   t[5058] := 0;
   t[5059] := 0;
   t[5060] := 0;
   t[5061] := 0;
   t[5062] := 0;
   t[5063] := 0;
   t[5064] := 0;
   t[5065] := 0;
   t[5066] := 0;
   t[5067] := 0;
   t[5068] := 0;
   t[5069] := 0;
   t[5070] := 0;
   t[5071] := 0;
   t[5072] := 0;
   t[5073] := 0;
   t[5074] := 0;
   t[5075] := 0;
   t[5076] := 0;
   t[5077] := 0;
   t[5078] := 0;
   t[5079] := 0;
   t[5080] := 0;
   t[5081] := 0;
   t[5082] := 0;
   t[5083] := 0;
   t[5084] := 0;
   t[5085] := 0;
   t[5086] := 0;
   t[5087] := 0;
   t[5088] := 0;
   t[5089] := 0;
   t[5090] := 0;
   t[5091] := 0;
   t[5092] := 0;
   t[5093] := 0;
   t[5094] := 0;
   t[5095] := 0;
   t[5096] := 0;
   t[5097] := 0;
   t[5098] := 0;
   t[5099] := 0;
   t[5100] := 0;
   t[5101] := 0;
   t[5102] := 0;
   t[5103] := 0;
   t[5104] := 0;
   t[5105] := 0;
   t[5106] := 0;
   t[5107] := 0;
   t[5108] := 0;
   t[5109] := 0;
   t[5110] := 0;
   t[5111] := 0;
   t[5112] := 0;
   t[5113] := 0;
   t[5114] := 0;
   t[5115] := 0;
   t[5116] := 0;
   t[5117] := 0;
   t[5118] := 0;
   t[5119] := 0;
   t[5120] := 0;
   t[5121] := 0;
   t[5122] := 0;
   t[5123] := 0;
   t[5124] := 0;
   t[5125] := 0;
   t[5126] := 0;
   t[5127] := 0;
   t[5128] := 0;
   t[5129] := 0;
   t[5130] := 0;
   t[5131] := 0;
   t[5132] := 0;
   t[5133] := 0;
   t[5134] := 0;
   t[5135] := 0;
   t[5136] := 0;
   t[5137] := 0;
   t[5138] := 0;
   t[5139] := 0;
   t[5140] := 0;
   t[5141] := 0;
   t[5142] := 0;
   t[5143] := 0;
   t[5144] := 0;
   t[5145] := 0;
   t[5146] := 0;
   t[5147] := 0;
   t[5148] := 0;
   t[5149] := 0;
   t[5150] := 0;
   t[5151] := 0;
   t[5152] := 0;
   t[5153] := 0;
   t[5154] := 0;
   t[5155] := 0;
   t[5156] := 0;
   t[5157] := 0;
   t[5158] := 0;
   t[5159] := 0;
   t[5160] := 0;
   t[5161] := 0;
   t[5162] := 0;
   t[5163] := 0;
   t[5164] := 0;
   t[5165] := 0;
   t[5166] := 0;
   t[5167] := 0;
   t[5168] := 0;
   t[5169] := 0;
   t[5170] := 0;
   t[5171] := 0;
   t[5172] := 0;
   t[5173] := 0;
   t[5174] := 0;
   t[5175] := 0;
   t[5176] := 0;
   t[5177] := 0;
   t[5178] := 0;
   t[5179] := 0;
   t[5180] := 0;
   t[5181] := 0;
   t[5182] := 0;
   t[5183] := 0;
   t[5184] := 0;
   t[5185] := 0;
   t[5186] := 0;
   t[5187] := 0;
   t[5188] := 0;
   t[5189] := 0;
   t[5190] := 0;
   t[5191] := 0;
   t[5192] := 0;
   t[5193] := 0;
   t[5194] := 0;
   t[5195] := 0;
   t[5196] := 0;
   t[5197] := 0;
   t[5198] := 0;
   t[5199] := 0;
   t[5200] := 0;
   t[5201] := 0;
   t[5202] := 0;
   t[5203] := 0;
   t[5204] := 0;
   t[5205] := 0;
   t[5206] := 0;
   t[5207] := 0;
   t[5208] := 0;
   t[5209] := 0;
   t[5210] := 0;
   t[5211] := 0;
   t[5212] := 0;
   t[5213] := 0;
   t[5214] := 0;
   t[5215] := 0;
   t[5216] := 0;
   t[5217] := 0;
   t[5218] := 0;
   t[5219] := 0;
   t[5220] := 0;
   t[5221] := 0;
   t[5222] := 0;
   t[5223] := 0;
   t[5224] := 0;
   t[5225] := 0;
   t[5226] := 0;
   t[5227] := 0;
   t[5228] := 0;
   t[5229] := 0;
   t[5230] := 0;
   t[5231] := 0;
   t[5232] := 0;
   t[5233] := 0;
   t[5234] := 0;
   t[5235] := 0;
   t[5236] := 0;
   t[5237] := 0;
   t[5238] := 0;
   t[5239] := 0;
   t[5240] := 0;
   t[5241] := 0;
   t[5242] := 0;
   t[5243] := 0;
   t[5244] := 0;
   t[5245] := 0;
   t[5246] := 0;
   t[5247] := 0;
   t[5248] := 0;
   t[5249] := 0;
   t[5250] := 0;
   t[5251] := 0;
   t[5252] := 0;
   t[5253] := 0;
   t[5254] := 0;
   t[5255] := 0;
   t[5256] := 0;
   t[5257] := 0;
   t[5258] := 0;
   t[5259] := 0;
   t[5260] := 0;
   t[5261] := 0;
   t[5262] := 0;
   t[5263] := 0;
   t[5264] := 0;
   t[5265] := 0;
   t[5266] := 0;
   t[5267] := 0;
   t[5268] := 0;
   t[5269] := 0;
   t[5270] := 0;
   t[5271] := 0;
   t[5272] := 0;
   t[5273] := 0;
   t[5274] := 0;
   t[5275] := 0;
   t[5276] := 0;
   t[5277] := 0;
   t[5278] := 0;
   t[5279] := 0;
   t[5280] := 0;
   t[5281] := 0;
   t[5282] := 0;
   t[5283] := 0;
   t[5284] := 0;
   t[5285] := 0;
   t[5286] := 0;
   t[5287] := 0;
   t[5288] := 0;
   t[5289] := 0;
   t[5290] := 0;
   t[5291] := 0;
   t[5292] := 0;
   t[5293] := 0;
   t[5294] := 0;
   t[5295] := 0;
   t[5296] := 0;
   t[5297] := 0;
   t[5298] := 0;
   t[5299] := 0;
   t[5300] := 0;
   t[5301] := 0;
   t[5302] := 0;
   t[5303] := 0;
   t[5304] := 0;
   t[5305] := 0;
   t[5306] := 0;
   t[5307] := 0;
   t[5308] := 0;
   t[5309] := 0;
   t[5310] := 0;
   t[5311] := 0;
   t[5312] := 0;
   t[5313] := 0;
   t[5314] := 0;
   t[5315] := 0;
   t[5316] := 0;
   t[5317] := 0;
   t[5318] := 0;
   t[5319] := 0;
   t[5320] := 0;
   t[5321] := 0;
   t[5322] := 0;
   t[5323] := 0;
   t[5324] := 0;
   t[5325] := 0;
   t[5326] := 0;
   t[5327] := 0;
   t[5328] := 0;
   t[5329] := 0;
   t[5330] := 0;
   t[5331] := 0;
   t[5332] := 0;
   t[5333] := 0;
   t[5334] := 0;
   t[5335] := 0;
   t[5336] := 0;
   t[5337] := 0;
   t[5338] := 0;
   t[5339] := 0;
   t[5340] := 0;
   t[5341] := 0;
   t[5342] := 0;
   t[5343] := 0;
   t[5344] := 0;
   t[5345] := 0;
   t[5346] := 0;
   t[5347] := 0;
   t[5348] := 0;
   t[5349] := 0;
   t[5350] := 0;
   t[5351] := 0;
   t[5352] := 0;
   t[5353] := 0;
   t[5354] := 0;
   t[5355] := 0;
   t[5356] := 0;
   t[5357] := 0;
   t[5358] := 0;
   t[5359] := 0;
   t[5360] := 0;
   t[5361] := 0;
   t[5362] := 0;
   t[5363] := 0;
   t[5364] := 0;
   t[5365] := 0;
   t[5366] := 0;
   t[5367] := 0;
   t[5368] := 0;
   t[5369] := 0;
   t[5370] := 0;
   t[5371] := 0;
   t[5372] := 0;
   t[5373] := 0;
   t[5374] := 0;
   t[5375] := 0;
   t[5376] := 0;
   t[5377] := 0;
   t[5378] := 0;
   t[5379] := 0;
   t[5380] := 0;
   t[5381] := 0;
   t[5382] := 0;
   t[5383] := 0;
   t[5384] := 0;
   t[5385] := 0;
   t[5386] := 0;
   t[5387] := 0;
   t[5388] := 0;
   t[5389] := 0;
   t[5390] := 0;
   t[5391] := 0;
   t[5392] := 0;
   t[5393] := 0;
   t[5394] := 0;
   t[5395] := 0;
   t[5396] := 0;
   t[5397] := 0;
   t[5398] := 0;
   t[5399] := 0;
   t[5400] := 0;
   t[5401] := 0;
   t[5402] := 0;
   t[5403] := 0;
   t[5404] := 0;
   t[5405] := 0;
   t[5406] := 0;
   t[5407] := 0;
   t[5408] := 0;
   t[5409] := 0;
   t[5410] := 0;
   t[5411] := 0;
   t[5412] := 0;
   t[5413] := 0;
   t[5414] := 0;
   t[5415] := 0;
   t[5416] := 0;
   t[5417] := 0;
   t[5418] := 0;
   t[5419] := 0;
   t[5420] := 0;
   t[5421] := 0;
   t[5422] := 0;
   t[5423] := 0;
   t[5424] := 0;
   t[5425] := 0;
   t[5426] := 0;
   t[5427] := 0;
   t[5428] := 0;
   t[5429] := 0;
   t[5430] := 0;
   t[5431] := 0;
   t[5432] := 0;
   t[5433] := 0;
   t[5434] := 0;
   t[5435] := 0;
   t[5436] := 0;
   t[5437] := 0;
   t[5438] := 0;
   t[5439] := 0;
   t[5440] := 0;
   t[5441] := 0;
   t[5442] := 0;
   t[5443] := 0;
   t[5444] := 0;
   t[5445] := 0;
   t[5446] := 0;
   t[5447] := 0;
   t[5448] := 0;
   t[5449] := 0;
   t[5450] := 0;
   t[5451] := 0;
   t[5452] := 0;
   t[5453] := 0;
   t[5454] := 0;
   t[5455] := 0;
   t[5456] := 0;
   t[5457] := 0;
   t[5458] := 0;
   t[5459] := 0;
   t[5460] := 0;
   t[5461] := 0;
   t[5462] := 0;
   t[5463] := 0;
   t[5464] := 0;
   t[5465] := 0;
   t[5466] := 0;
   t[5467] := 0;
   t[5468] := 0;
   t[5469] := 0;
   t[5470] := 0;
   t[5471] := 0;
   t[5472] := 0;
   t[5473] := 0;
   t[5474] := 0;
   t[5475] := 0;
   t[5476] := 0;
   t[5477] := 0;
   t[5478] := 0;
   t[5479] := 0;
   t[5480] := 0;
   t[5481] := 0;
   t[5482] := 0;
   t[5483] := 0;
   t[5484] := 0;
   t[5485] := 0;
   t[5486] := 0;
   t[5487] := 0;
   t[5488] := 0;
   t[5489] := 0;
   t[5490] := 0;
   t[5491] := 0;
   t[5492] := 0;
   t[5493] := 0;
   t[5494] := 0;
   t[5495] := 0;
   t[5496] := 0;
   t[5497] := 0;
   t[5498] := 0;
   t[5499] := 0;
   t[5500] := 0;
   t[5501] := 0;
   t[5502] := 0;
   t[5503] := 0;
   t[5504] := 0;
   t[5505] := 0;
   t[5506] := 0;
   t[5507] := 0;
   t[5508] := 0;
   t[5509] := 0;
   t[5510] := 0;
   t[5511] := 0;
   t[5512] := 0;
   t[5513] := 0;
   t[5514] := 0;
   t[5515] := 0;
   t[5516] := 0;
   t[5517] := 0;
   t[5518] := 0;
   t[5519] := 0;
   t[5520] := 0;
   t[5521] := 0;
   t[5522] := 0;
   t[5523] := 0;
   t[5524] := 0;
   t[5525] := 0;
   t[5526] := 0;
   t[5527] := 0;
   t[5528] := 0;
   t[5529] := 0;
   t[5530] := 0;
   t[5531] := 0;
   t[5532] := 0;
   t[5533] := 0;
   t[5534] := 0;
   t[5535] := 0;
   t[5536] := 0;
   t[5537] := 0;
   t[5538] := 0;
   t[5539] := 0;
   t[5540] := 0;
   t[5541] := 0;
   t[5542] := 0;
   t[5543] := 0;
   t[5544] := 0;
   t[5545] := 0;
   t[5546] := 0;
   t[5547] := 0;
   t[5548] := 0;
   t[5549] := 0;
   t[5550] := 0;
   t[5551] := 0;
   t[5552] := 0;
   t[5553] := 0;
   t[5554] := 0;
   t[5555] := 0;
   t[5556] := 0;
   t[5557] := 0;
   t[5558] := 0;
   t[5559] := 0;
   t[5560] := 0;
   t[5561] := 0;
   t[5562] := 0;
   t[5563] := 0;
   t[5564] := 0;
   t[5565] := 0;
   t[5566] := 0;
   t[5567] := 0;
   t[5568] := 0;
   t[5569] := 0;
   t[5570] := 0;
   t[5571] := 0;
   t[5572] := 0;
   t[5573] := 0;
   t[5574] := 0;
   t[5575] := 0;
   t[5576] := 0;
   t[5577] := 0;
   t[5578] := 0;
   t[5579] := 0;
   t[5580] := 0;
   t[5581] := 0;
   t[5582] := 0;
   t[5583] := 0;
   t[5584] := 0;
   t[5585] := 0;
   t[5586] := 0;
   t[5587] := 0;
   t[5588] := 0;
   t[5589] := 0;
   t[5590] := 0;
   t[5591] := 0;
   t[5592] := 0;
   t[5593] := 0;
   t[5594] := 0;
   t[5595] := 0;
   t[5596] := 0;
   t[5597] := 0;
   t[5598] := 0;
   t[5599] := 0;
   t[5600] := 0;
   t[5601] := 0;
   t[5602] := 0;
   t[5603] := 0;
   t[5604] := 0;
   t[5605] := 0;
   t[5606] := 0;
   t[5607] := 0;
   t[5608] := 0;
   t[5609] := 0;
   t[5610] := 0;
   t[5611] := 0;
   t[5612] := 0;
   t[5613] := 0;
   t[5614] := 0;
   t[5615] := 0;
   t[5616] := 0;
   t[5617] := 0;
   t[5618] := 0;
   t[5619] := 0;
   t[5620] := 0;
   t[5621] := 0;
   t[5622] := 0;
   t[5623] := 0;
   t[5624] := 0;
   t[5625] := 0;
   t[5626] := 0;
   t[5627] := 0;
   t[5628] := 0;
   t[5629] := 0;
   t[5630] := 0;
   t[5631] := 0;
   t[5632] := 0;
   t[5633] := 0;
   t[5634] := 0;
   t[5635] := 0;
   t[5636] := 0;
   t[5637] := 0;
   t[5638] := 0;
   t[5639] := 0;
   t[5640] := 0;
   t[5641] := 0;
   t[5642] := 0;
   t[5643] := 0;
   t[5644] := 0;
   t[5645] := 0;
   t[5646] := 0;
   t[5647] := 0;
   t[5648] := 0;
   t[5649] := 0;
   t[5650] := 0;
   t[5651] := 0;
   t[5652] := 0;
   t[5653] := 0;
   t[5654] := 0;
   t[5655] := 0;
   t[5656] := 0;
   t[5657] := 0;
   t[5658] := 0;
   t[5659] := 0;
   t[5660] := 0;
   t[5661] := 0;
   t[5662] := 0;
   t[5663] := 0;
   t[5664] := 0;
   t[5665] := 0;
   t[5666] := 0;
   t[5667] := 0;
   t[5668] := 0;
   t[5669] := 0;
   t[5670] := 0;
   t[5671] := 0;
   t[5672] := 0;
   t[5673] := 0;
   t[5674] := 0;
   t[5675] := 0;
   t[5676] := 0;
   t[5677] := 0;
   t[5678] := 0;
   t[5679] := 0;
   t[5680] := 0;
   t[5681] := 0;
   t[5682] := 0;
   t[5683] := 0;
   t[5684] := 0;
   t[5685] := 0;
   t[5686] := 0;
   t[5687] := 0;
   t[5688] := 0;
   t[5689] := 0;
   t[5690] := 0;
   t[5691] := 0;
   t[5692] := 0;
   t[5693] := 0;
   t[5694] := 0;
   t[5695] := 0;
   t[5696] := 0;
   t[5697] := 0;
   t[5698] := 0;
   t[5699] := 0;
   t[5700] := 0;
   t[5701] := 0;
   t[5702] := 0;
   t[5703] := 0;
   t[5704] := 0;
   t[5705] := 0;
   t[5706] := 0;
   t[5707] := 0;
   t[5708] := 0;
   t[5709] := 0;
   t[5710] := 0;
   t[5711] := 0;
   t[5712] := 0;
   t[5713] := 0;
   t[5714] := 0;
   t[5715] := 0;
   t[5716] := 0;
   t[5717] := 0;
   t[5718] := 0;
   t[5719] := 0;
   t[5720] := 0;
   t[5721] := 0;
   t[5722] := 0;
   t[5723] := 0;
   t[5724] := 0;
   t[5725] := 0;
   t[5726] := 0;
   t[5727] := 0;
   t[5728] := 0;
   t[5729] := 0;
   t[5730] := 0;
   t[5731] := 0;
   t[5732] := 0;
   t[5733] := 0;
   t[5734] := 0;
   t[5735] := 0;
   t[5736] := 0;
   t[5737] := 0;
   t[5738] := 0;
   t[5739] := 0;
   t[5740] := 0;
   t[5741] := 0;
   t[5742] := 0;
   t[5743] := 0;
   t[5744] := 0;
   t[5745] := 0;
   t[5746] := 0;
   t[5747] := 0;
   t[5748] := 0;
   t[5749] := 0;
   t[5750] := 0;
   t[5751] := 0;
   t[5752] := 0;
   t[5753] := 0;
   t[5754] := 0;
   t[5755] := 0;
   t[5756] := 0;
   t[5757] := 0;
   t[5758] := 0;
   t[5759] := 0;
   t[5760] := 0;
   t[5761] := 0;
   t[5762] := 0;
   t[5763] := 0;
   t[5764] := 0;
   t[5765] := 0;
   t[5766] := 0;
   t[5767] := 0;
   t[5768] := 0;
   t[5769] := 0;
   t[5770] := 0;
   t[5771] := 0;
   t[5772] := 0;
   t[5773] := 0;
   t[5774] := 0;
   t[5775] := 0;
   t[5776] := 0;
   t[5777] := 0;
   t[5778] := 0;
   t[5779] := 0;
   t[5780] := 0;
   t[5781] := 0;
   t[5782] := 0;
   t[5783] := 0;
   t[5784] := 0;
   t[5785] := 0;
   t[5786] := 0;
   t[5787] := 0;
   t[5788] := 0;
   t[5789] := 0;
   t[5790] := 0;
   t[5791] := 0;
   t[5792] := 0;
   t[5793] := 0;
   t[5794] := 0;
   t[5795] := 0;
   t[5796] := 0;
   t[5797] := 0;
   t[5798] := 0;
   t[5799] := 0;
   t[5800] := 0;
   t[5801] := 0;
   t[5802] := 0;
   t[5803] := 0;
   t[5804] := 0;
   t[5805] := 0;
   t[5806] := 0;
   t[5807] := 0;
   t[5808] := 0;
   t[5809] := 0;
   t[5810] := 0;
   t[5811] := 0;
   t[5812] := 0;
   t[5813] := 0;
   t[5814] := 0;
   t[5815] := 0;
   t[5816] := 0;
   t[5817] := 0;
   t[5818] := 0;
   t[5819] := 0;
   t[5820] := 0;
   t[5821] := 0;
   t[5822] := 0;
   t[5823] := 0;
   t[5824] := 0;
   t[5825] := 0;
   t[5826] := 0;
   t[5827] := 0;
   t[5828] := 0;
   t[5829] := 0;
   t[5830] := 0;
   t[5831] := 0;
   t[5832] := 0;
   t[5833] := 0;
   t[5834] := 0;
   t[5835] := 0;
   t[5836] := 0;
   t[5837] := 0;
   t[5838] := 0;
   t[5839] := 0;
   t[5840] := 0;
   t[5841] := 0;
   t[5842] := 0;
   t[5843] := 0;
   t[5844] := 0;
   t[5845] := 0;
   t[5846] := 0;
   t[5847] := 0;
   t[5848] := 0;
   t[5849] := 0;
   t[5850] := 0;
   t[5851] := 0;
   t[5852] := 0;
   t[5853] := 0;
   t[5854] := 0;
   t[5855] := 0;
   t[5856] := 0;
   t[5857] := 0;
   t[5858] := 0;
   t[5859] := 0;
   t[5860] := 0;
   t[5861] := 0;
   t[5862] := 0;
   t[5863] := 0;
   t[5864] := 0;
   t[5865] := 0;
   t[5866] := 0;
   t[5867] := 0;
   t[5868] := 0;
   t[5869] := 0;
   t[5870] := 0;
   t[5871] := 0;
   t[5872] := 0;
   t[5873] := 0;
   t[5874] := 0;
   t[5875] := 0;
   t[5876] := 0;
   t[5877] := 0;
   t[5878] := 0;
   t[5879] := 0;
   t[5880] := 0;
   t[5881] := 0;
   t[5882] := 0;
   t[5883] := 0;
   t[5884] := 0;
   t[5885] := 0;
   t[5886] := 0;
   t[5887] := 0;
   t[5888] := 0;
   t[5889] := 0;
   t[5890] := 0;
   t[5891] := 0;
   t[5892] := 0;
   t[5893] := 0;
   t[5894] := 0;
   t[5895] := 0;
   t[5896] := 0;
   t[5897] := 0;
   t[5898] := 0;
   t[5899] := 0;
   t[5900] := 0;
   t[5901] := 0;
   t[5902] := 0;
   t[5903] := 0;
   t[5904] := 0;
   t[5905] := 0;
   t[5906] := 0;
   t[5907] := 0;
   t[5908] := 0;
   t[5909] := 0;
   t[5910] := 0;
   t[5911] := 0;
   t[5912] := 0;
   t[5913] := 0;
   t[5914] := 0;
   t[5915] := 0;
   t[5916] := 0;
   t[5917] := 0;
   t[5918] := 0;
   t[5919] := 0;
   t[5920] := 0;
   t[5921] := 0;
   t[5922] := 0;
   t[5923] := 0;
   t[5924] := 0;
   t[5925] := 0;
   t[5926] := 0;
   t[5927] := 0;
   t[5928] := 0;
   t[5929] := 0;
   t[5930] := 0;
   t[5931] := 0;
   t[5932] := 0;
   t[5933] := 0;
   t[5934] := 0;
   t[5935] := 0;
   t[5936] := 0;
   t[5937] := 0;
   t[5938] := 0;
   t[5939] := 0;
   t[5940] := 0;
   t[5941] := 0;
   t[5942] := 0;
   t[5943] := 0;
   t[5944] := 0;
   t[5945] := 0;
   t[5946] := 0;
   t[5947] := 0;
   t[5948] := 0;
   t[5949] := 0;
   t[5950] := 0;
   t[5951] := 0;
   t[5952] := 0;
   t[5953] := 0;
   t[5954] := 0;
   t[5955] := 0;
   t[5956] := 0;
   t[5957] := 0;
   t[5958] := 0;
   t[5959] := 0;
   t[5960] := 0;
   t[5961] := 0;
   t[5962] := 0;
   t[5963] := 0;
   t[5964] := 0;
   t[5965] := 0;
   t[5966] := 0;
   t[5967] := 0;
   t[5968] := 0;
   t[5969] := 0;
   t[5970] := 0;
   t[5971] := 0;
   t[5972] := 0;
   t[5973] := 0;
   t[5974] := 0;
   t[5975] := 0;
   t[5976] := 0;
   t[5977] := 0;
   t[5978] := 0;
   t[5979] := 0;
   t[5980] := 0;
   t[5981] := 0;
   t[5982] := 0;
   t[5983] := 0;
   t[5984] := 0;
   t[5985] := 0;
   t[5986] := 0;
   t[5987] := 0;
   t[5988] := 0;
   t[5989] := 0;
   t[5990] := 0;
   t[5991] := 0;
   t[5992] := 0;
   t[5993] := 0;
   t[5994] := 0;
   t[5995] := 0;
   t[5996] := 0;
   t[5997] := 0;
   t[5998] := 0;
   t[5999] := 0;
   t[6000] := 0;
   t[6001] := 0;
   t[6002] := 0;
   t[6003] := 0;
   t[6004] := 0;
   t[6005] := 0;
   t[6006] := 0;
   t[6007] := 0;
   t[6008] := 0;
   t[6009] := 0;
   t[6010] := 0;
   t[6011] := 0;
   t[6012] := 0;
   t[6013] := 0;
   t[6014] := 0;
   t[6015] := 0;
   t[6016] := 0;
   t[6017] := 0;
   t[6018] := 0;
   t[6019] := 0;
   t[6020] := 0;
   t[6021] := 0;
   t[6022] := 0;
   t[6023] := 0;
   t[6024] := 0;
   t[6025] := 0;
   t[6026] := 0;
   t[6027] := 0;
   t[6028] := 0;
   t[6029] := 0;
   t[6030] := 0;
   t[6031] := 0;
   t[6032] := 0;
   t[6033] := 0;
   t[6034] := 0;
   t[6035] := 0;
   t[6036] := 0;
   t[6037] := 0;
   t[6038] := 0;
   t[6039] := 0;
   t[6040] := 0;
   t[6041] := 0;
   t[6042] := 0;
   t[6043] := 0;
   t[6044] := 0;
   t[6045] := 0;
   t[6046] := 0;
   t[6047] := 0;
   t[6048] := 0;
   t[6049] := 0;
   t[6050] := 0;
   t[6051] := 0;
   t[6052] := 0;
   t[6053] := 0;
   t[6054] := 0;
   t[6055] := 0;
   t[6056] := 0;
   t[6057] := 0;
   t[6058] := 0;
   t[6059] := 0;
   t[6060] := 0;
   t[6061] := 0;
   t[6062] := 0;
   t[6063] := 0;
   t[6064] := 0;
   t[6065] := 0;
   t[6066] := 0;
   t[6067] := 0;
   t[6068] := 0;
   t[6069] := 0;
   t[6070] := 0;
   t[6071] := 0;
   t[6072] := 0;
   t[6073] := 0;
   t[6074] := 0;
   t[6075] := 0;
   t[6076] := 0;
   t[6077] := 0;
   t[6078] := 0;
   t[6079] := 0;
   t[6080] := 0;
   t[6081] := 0;
   t[6082] := 0;
   t[6083] := 0;
   t[6084] := 0;
   t[6085] := 0;
   t[6086] := 0;
   t[6087] := 0;
   t[6088] := 0;
   t[6089] := 0;
   t[6090] := 0;
   t[6091] := 0;
   t[6092] := 0;
   t[6093] := 0;
   t[6094] := 0;
   t[6095] := 0;
   t[6096] := 0;
   t[6097] := 0;
   t[6098] := 0;
   t[6099] := 0;
   t[6100] := 0;
   t[6101] := 0;
   t[6102] := 0;
   t[6103] := 0;
   t[6104] := 0;
   t[6105] := 0;
   t[6106] := 0;
   t[6107] := 0;
   t[6108] := 0;
   t[6109] := 0;
   t[6110] := 0;
   t[6111] := 0;
   t[6112] := 0;
   t[6113] := 0;
   t[6114] := 0;
   t[6115] := 0;
   t[6116] := 0;
   t[6117] := 0;
   t[6118] := 0;
   t[6119] := 0;
   t[6120] := 0;
   t[6121] := 0;
   t[6122] := 0;
   t[6123] := 0;
   t[6124] := 0;
   t[6125] := 0;
   t[6126] := 0;
   t[6127] := 0;
   t[6128] := 0;
   t[6129] := 0;
   t[6130] := 0;
   t[6131] := 0;
   t[6132] := 0;
   t[6133] := 0;
   t[6134] := 0;
   t[6135] := 0;
   t[6136] := 0;
   t[6137] := 0;
   t[6138] := 0;
   t[6139] := 0;
   t[6140] := 0;
   t[6141] := 0;
   t[6142] := 0;
   t[6143] := 0;
   t[6144] := 0;
   t[6145] := 0;
   t[6146] := 0;
   t[6147] := 0;
   t[6148] := 0;
   t[6149] := 0;
   t[6150] := 0;
   t[6151] := 0;
   t[6152] := 0;
   t[6153] := 0;
   t[6154] := 0;
   t[6155] := 0;
   t[6156] := 0;
   t[6157] := 0;
   t[6158] := 0;
   t[6159] := 0;
   t[6160] := 0;
   t[6161] := 0;
   t[6162] := 0;
   t[6163] := 0;
   t[6164] := 0;
   t[6165] := 0;
   t[6166] := 0;
   t[6167] := 0;
   t[6168] := 0;
   t[6169] := 0;
   t[6170] := 0;
   t[6171] := 0;
   t[6172] := 0;
   t[6173] := 0;
   t[6174] := 0;
   t[6175] := 0;
   t[6176] := 0;
   t[6177] := 0;
   t[6178] := 0;
   t[6179] := 0;
   t[6180] := 0;
   t[6181] := 0;
   t[6182] := 0;
   t[6183] := 0;
   t[6184] := 0;
   t[6185] := 0;
   t[6186] := 0;
   t[6187] := 0;
   t[6188] := 0;
   t[6189] := 0;
   t[6190] := 0;
   t[6191] := 0;
   t[6192] := 0;
   t[6193] := 0;
   t[6194] := 0;
   t[6195] := 0;
   t[6196] := 0;
   t[6197] := 0;
   t[6198] := 0;
   t[6199] := 0;
   t[6200] := 0;
   t[6201] := 0;
   t[6202] := 0;
   t[6203] := 0;
   t[6204] := 0;
   t[6205] := 0;
   t[6206] := 0;
   t[6207] := 0;
   t[6208] := 0;
   t[6209] := 0;
   t[6210] := 0;
   t[6211] := 0;
   t[6212] := 0;
   t[6213] := 0;
   t[6214] := 0;
   t[6215] := 0;
   t[6216] := 0;
   t[6217] := 0;
   t[6218] := 0;
   t[6219] := 0;
   t[6220] := 0;
   t[6221] := 0;
   t[6222] := 0;
   t[6223] := 0;
   t[6224] := 0;
   t[6225] := 0;
   t[6226] := 0;
   t[6227] := 0;
   t[6228] := 0;
   t[6229] := 0;
   t[6230] := 0;
   t[6231] := 0;
   t[6232] := 0;
   t[6233] := 0;
   t[6234] := 0;
   t[6235] := 0;
   t[6236] := 0;
   t[6237] := 0;
   t[6238] := 0;
   t[6239] := 0;
   t[6240] := 0;
   t[6241] := 0;
   t[6242] := 0;
   t[6243] := 0;
   t[6244] := 0;
   t[6245] := 0;
   t[6246] := 0;
   t[6247] := 0;
   t[6248] := 0;
   t[6249] := 0;
   t[6250] := 0;
   t[6251] := 0;
   t[6252] := 0;
   t[6253] := 0;
   t[6254] := 0;
   t[6255] := 0;
   t[6256] := 0;
   t[6257] := 0;
   t[6258] := 0;
   t[6259] := 0;
   t[6260] := 0;
   t[6261] := 0;
   t[6262] := 0;
   t[6263] := 0;
   t[6264] := 0;
   t[6265] := 0;
   t[6266] := 0;
   t[6267] := 0;
   t[6268] := 0;
   t[6269] := 0;
   t[6270] := 0;
   t[6271] := 0;
   t[6272] := 0;
   t[6273] := 0;
   t[6274] := 0;
   t[6275] := 0;
   t[6276] := 0;
   t[6277] := 0;
   t[6278] := 0;
   t[6279] := 0;
   t[6280] := 0;
   t[6281] := 0;
   t[6282] := 0;
   t[6283] := 0;
   t[6284] := 0;
   t[6285] := 0;
   t[6286] := 0;
   t[6287] := 0;
   t[6288] := 0;
   t[6289] := 0;
   t[6290] := 0;
   t[6291] := 0;
   t[6292] := 0;
   t[6293] := 0;
   t[6294] := 0;
   t[6295] := 0;
   t[6296] := 0;
   t[6297] := 0;
   t[6298] := 0;
   t[6299] := 0;
   t[6300] := 0;
   t[6301] := 0;
   t[6302] := 0;
   t[6303] := 0;
   t[6304] := 0;
   t[6305] := 0;
   t[6306] := 0;
   t[6307] := 0;
   t[6308] := 0;
   t[6309] := 0;
   t[6310] := 0;
   t[6311] := 0;
   t[6312] := 0;
   t[6313] := 0;
   t[6314] := 0;
   t[6315] := 0;
   t[6316] := 0;
   t[6317] := 0;
   t[6318] := 0;
   t[6319] := 0;
   t[6320] := 0;
   t[6321] := 0;
   t[6322] := 0;
   t[6323] := 0;
   t[6324] := 0;
   t[6325] := 0;
   t[6326] := 0;
   t[6327] := 0;
   t[6328] := 0;
   t[6329] := 0;
   t[6330] := 0;
   t[6331] := 0;
   t[6332] := 0;
   t[6333] := 0;
   t[6334] := 0;
   t[6335] := 0;
   t[6336] := 0;
   t[6337] := 0;
   t[6338] := 0;
   t[6339] := 0;
   t[6340] := 0;
   t[6341] := 0;
   t[6342] := 0;
   t[6343] := 0;
   t[6344] := 0;
   t[6345] := 0;
   t[6346] := 0;
   t[6347] := 0;
   t[6348] := 0;
   t[6349] := 0;
   t[6350] := 0;
   t[6351] := 0;
   t[6352] := 0;
   t[6353] := 0;
   t[6354] := 0;
   t[6355] := 0;
   t[6356] := 0;
   t[6357] := 0;
   t[6358] := 0;
   t[6359] := 0;
   t[6360] := 0;
   t[6361] := 0;
   t[6362] := 0;
   t[6363] := 0;
   t[6364] := 0;
   t[6365] := 0;
   t[6366] := 0;
   t[6367] := 0;
   t[6368] := 0;
   t[6369] := 0;
   t[6370] := 0;
   t[6371] := 0;
   t[6372] := 0;
   t[6373] := 0;
   t[6374] := 0;
   t[6375] := 0;
   t[6376] := 0;
   t[6377] := 0;
   t[6378] := 0;
   t[6379] := 0;
   t[6380] := 0;
   t[6381] := 0;
   t[6382] := 0;
   t[6383] := 0;
   t[6384] := 0;
   t[6385] := 0;
   t[6386] := 0;
   t[6387] := 0;
   t[6388] := 0;
   t[6389] := 0;
   t[6390] := 0;
   t[6391] := 0;
   t[6392] := 0;
   t[6393] := 0;
   t[6394] := 0;
   t[6395] := 0;
   t[6396] := 0;
   t[6397] := 0;
   t[6398] := 0;
   t[6399] := 0;
   t[6400] := 0;
   t[6401] := 0;
   t[6402] := 0;
   t[6403] := 0;
   t[6404] := 0;
   t[6405] := 0;
   t[6406] := 0;
   t[6407] := 0;
   t[6408] := 0;
   t[6409] := 0;
   t[6410] := 0;
   t[6411] := 0;
   t[6412] := 0;
   t[6413] := 0;
   t[6414] := 0;
   t[6415] := 0;
   t[6416] := 0;
   t[6417] := 0;
   t[6418] := 0;
   t[6419] := 0;
   t[6420] := 0;
   t[6421] := 0;
   t[6422] := 0;
   t[6423] := 0;
   t[6424] := 0;
   t[6425] := 0;
   t[6426] := 0;
   t[6427] := 0;
   t[6428] := 0;
   t[6429] := 0;
   t[6430] := 0;
   t[6431] := 0;
   t[6432] := 0;
   t[6433] := 0;
   t[6434] := 0;
   t[6435] := 0;
   t[6436] := 0;
   t[6437] := 0;
   t[6438] := 0;
   t[6439] := 0;
   t[6440] := 0;
   t[6441] := 0;
   t[6442] := 0;
   t[6443] := 0;
   t[6444] := 0;
   t[6445] := 0;
   t[6446] := 0;
   t[6447] := 0;
   t[6448] := 0;
   t[6449] := 0;
   t[6450] := 0;
   t[6451] := 0;
   t[6452] := 0;
   t[6453] := 0;
   t[6454] := 0;
   t[6455] := 0;
   t[6456] := 0;
   t[6457] := 0;
   t[6458] := 0;
   t[6459] := 0;
   t[6460] := 0;
   t[6461] := 0;
   t[6462] := 0;
   t[6463] := 0;
   t[6464] := 0;
   t[6465] := 0;
   t[6466] := 0;
   t[6467] := 0;
   t[6468] := 0;
   t[6469] := 0;
   t[6470] := 0;
   t[6471] := 0;
   t[6472] := 0;
   t[6473] := 0;
   t[6474] := 0;
   t[6475] := 0;
   t[6476] := 0;
   t[6477] := 0;
   t[6478] := 0;
   t[6479] := 0;
   t[6480] := 0;
   t[6481] := 0;
   t[6482] := 0;
   t[6483] := 0;
   t[6484] := 0;
   t[6485] := 0;
   t[6486] := 0;
   t[6487] := 0;
   t[6488] := 0;
   t[6489] := 0;
   t[6490] := 0;
   t[6491] := 0;
   t[6492] := 0;
   t[6493] := 0;
   t[6494] := 0;
   t[6495] := 0;
   t[6496] := 0;
   t[6497] := 0;
   t[6498] := 0;
   t[6499] := 0;
   t[6500] := 0;
   t[6501] := 0;
   t[6502] := 0;
   t[6503] := 0;
   t[6504] := 0;
   t[6505] := 0;
   t[6506] := 0;
   t[6507] := 0;
   t[6508] := 0;
   t[6509] := 0;
   t[6510] := 0;
   t[6511] := 0;
   t[6512] := 0;
   t[6513] := 0;
   t[6514] := 0;
   t[6515] := 0;
   t[6516] := 0;
   t[6517] := 0;
   t[6518] := 0;
   t[6519] := 0;
   t[6520] := 0;
   t[6521] := 0;
   t[6522] := 0;
   t[6523] := 0;
   t[6524] := 0;
   t[6525] := 0;
   t[6526] := 0;
   t[6527] := 0;
   t[6528] := 0;
   t[6529] := 0;
   t[6530] := 0;
   t[6531] := 0;
   t[6532] := 0;
   t[6533] := 0;
   t[6534] := 0;
   t[6535] := 0;
   t[6536] := 0;
   t[6537] := 0;
   t[6538] := 0;
   t[6539] := 0;
   t[6540] := 0;
   t[6541] := 0;
   t[6542] := 0;
   t[6543] := 0;
   t[6544] := 0;
   t[6545] := 0;
   t[6546] := 0;
   t[6547] := 0;
   t[6548] := 0;
   t[6549] := 0;
   t[6550] := 0;
   t[6551] := 0;
   t[6552] := 0;
   t[6553] := 0;
   t[6554] := 0;
   t[6555] := 0;
   t[6556] := 0;
   t[6557] := 0;
   t[6558] := 0;
   t[6559] := 0;
   t[6560] := 0;
   t[6561] := 0;
   t[6562] := 0;
   t[6563] := 0;
   t[6564] := 0;
   t[6565] := 0;
   t[6566] := 0;
   t[6567] := 0;
   t[6568] := 0;
   t[6569] := 0;
   t[6570] := 0;
   t[6571] := 0;
   t[6572] := 0;
   t[6573] := 0;
   t[6574] := 0;
   t[6575] := 0;
   t[6576] := 0;
   t[6577] := 0;
   t[6578] := 0;
   t[6579] := 0;
   t[6580] := 0;
   t[6581] := 0;
   t[6582] := 0;
   t[6583] := 0;
   t[6584] := 0;
   t[6585] := 0;
   t[6586] := 0;
   t[6587] := 0;
   t[6588] := 0;
   t[6589] := 0;
   t[6590] := 0;
   t[6591] := 0;
   t[6592] := 0;
   t[6593] := 0;
   t[6594] := 0;
   t[6595] := 0;
   t[6596] := 0;
   t[6597] := 0;
   t[6598] := 0;
   t[6599] := 0;
   t[6600] := 0;
   t[6601] := 0;
   t[6602] := 0;
   t[6603] := 0;
   t[6604] := 0;
   t[6605] := 0;
   t[6606] := 0;
   t[6607] := 0;
   t[6608] := 0;
   t[6609] := 0;
   t[6610] := 0;
   t[6611] := 0;
   t[6612] := 0;
   t[6613] := 0;
   t[6614] := 0;
   t[6615] := 0;
   t[6616] := 0;
   t[6617] := 0;
   t[6618] := 0;
   t[6619] := 0;
   t[6620] := 0;
   t[6621] := 0;
   t[6622] := 0;
   t[6623] := 0;
   t[6624] := 0;
   t[6625] := 0;
   t[6626] := 0;
   t[6627] := 0;
   t[6628] := 0;
   t[6629] := 0;
   t[6630] := 0;
   t[6631] := 0;
   t[6632] := 0;
   t[6633] := 0;
   t[6634] := 0;
   t[6635] := 0;
   t[6636] := 0;
   t[6637] := 0;
   t[6638] := 0;
   t[6639] := 0;
   t[6640] := 0;
   t[6641] := 0;
   t[6642] := 0;
   t[6643] := 0;
   t[6644] := 0;
   t[6645] := 0;
   t[6646] := 0;
   t[6647] := 0;
   t[6648] := 0;
   t[6649] := 0;
   t[6650] := 0;
   t[6651] := 0;
   t[6652] := 0;
   t[6653] := 0;
   t[6654] := 0;
   t[6655] := 0;
   t[6656] := 0;
   t[6657] := 0;
   t[6658] := 0;
   t[6659] := 0;
   t[6660] := 0;
   t[6661] := 0;
   t[6662] := 0;
   t[6663] := 0;
   t[6664] := 0;
   t[6665] := 0;
   t[6666] := 0;
   t[6667] := 0;
   t[6668] := 0;
   t[6669] := 0;
   t[6670] := 0;
   t[6671] := 0;
   t[6672] := 0;
   t[6673] := 0;
   t[6674] := 0;
   t[6675] := 0;
   t[6676] := 0;
   t[6677] := 0;
   t[6678] := 0;
   t[6679] := 0;
   t[6680] := 0;
   t[6681] := 0;
   t[6682] := 0;
   t[6683] := 0;
   t[6684] := 0;
   t[6685] := 0;
   t[6686] := 0;
   t[6687] := 0;
   t[6688] := 0;
   t[6689] := 0;
   t[6690] := 0;
   t[6691] := 0;
   t[6692] := 0;
   t[6693] := 0;
   t[6694] := 0;
   t[6695] := 0;
   t[6696] := 0;
   t[6697] := 0;
   t[6698] := 0;
   t[6699] := 0;
   t[6700] := 0;
   t[6701] := 0;
   t[6702] := 0;
   t[6703] := 0;
   t[6704] := 0;
   t[6705] := 0;
   t[6706] := 0;
   t[6707] := 0;
   t[6708] := 0;
   t[6709] := 0;
   t[6710] := 0;
   t[6711] := 0;
   t[6712] := 0;
   t[6713] := 0;
   t[6714] := 0;
   t[6715] := 0;
   t[6716] := 0;
   t[6717] := 0;
   t[6718] := 0;
   t[6719] := 0;
   t[6720] := 0;
   t[6721] := 0;
   t[6722] := 0;
   t[6723] := 0;
   t[6724] := 0;
   t[6725] := 0;
   t[6726] := 0;
   t[6727] := 0;
   t[6728] := 0;
   t[6729] := 0;
   t[6730] := 0;
   t[6731] := 0;
   t[6732] := 0;
   t[6733] := 0;
   t[6734] := 0;
   t[6735] := 0;
   t[6736] := 0;
   t[6737] := 0;
   t[6738] := 0;
   t[6739] := 0;
   t[6740] := 0;
   t[6741] := 0;
   t[6742] := 0;
   t[6743] := 0;
   t[6744] := 0;
   t[6745] := 0;
   t[6746] := 0;
   t[6747] := 0;
   t[6748] := 0;
   t[6749] := 0;
   t[6750] := 0;
   t[6751] := 0;
   t[6752] := 0;
   t[6753] := 0;
   t[6754] := 0;
   t[6755] := 0;
   t[6756] := 0;
   t[6757] := 0;
   t[6758] := 0;
   t[6759] := 0;
   t[6760] := 0;
   t[6761] := 0;
   t[6762] := 0;
   t[6763] := 0;
   t[6764] := 0;
   t[6765] := 0;
   t[6766] := 0;
   t[6767] := 0;
   t[6768] := 0;
   t[6769] := 0;
   t[6770] := 0;
   t[6771] := 0;
   t[6772] := 0;
   t[6773] := 0;
   t[6774] := 0;
   t[6775] := 0;
   t[6776] := 0;
   t[6777] := 0;
   t[6778] := 0;
   t[6779] := 0;
   t[6780] := 0;
   t[6781] := 0;
   t[6782] := 0;
   t[6783] := 0;
   t[6784] := 0;
   t[6785] := 0;
   t[6786] := 0;
   t[6787] := 0;
   t[6788] := 0;
   t[6789] := 0;
   t[6790] := 0;
   t[6791] := 0;
   t[6792] := 0;
   t[6793] := 0;
   t[6794] := 0;
   t[6795] := 0;
   t[6796] := 0;
   t[6797] := 0;
   t[6798] := 0;
   t[6799] := 0;
   t[6800] := 0;
   t[6801] := 0;
   t[6802] := 0;
   t[6803] := 0;
   t[6804] := 0;
   t[6805] := 0;
   t[6806] := 0;
   t[6807] := 0;
   t[6808] := 0;
   t[6809] := 0;
   t[6810] := 0;
   t[6811] := 0;
   t[6812] := 0;
   t[6813] := 0;
   t[6814] := 0;
   t[6815] := 0;
   t[6816] := 0;
   t[6817] := 0;
   t[6818] := 0;
   t[6819] := 0;
   t[6820] := 0;
   t[6821] := 0;
   t[6822] := 0;
   t[6823] := 0;
   t[6824] := 0;
   t[6825] := 0;
   t[6826] := 0;
   t[6827] := 0;
   t[6828] := 0;
   t[6829] := 0;
   t[6830] := 0;
   t[6831] := 0;
   t[6832] := 0;
   t[6833] := 0;
   t[6834] := 0;
   t[6835] := 0;
   t[6836] := 0;
   t[6837] := 0;
   t[6838] := 0;
   t[6839] := 0;
   t[6840] := 0;
   t[6841] := 0;
   t[6842] := 0;
   t[6843] := 0;
   t[6844] := 0;
   t[6845] := 0;
   t[6846] := 0;
   t[6847] := 0;
   t[6848] := 0;
   t[6849] := 0;
   t[6850] := 0;
   t[6851] := 0;
   t[6852] := 0;
   t[6853] := 0;
   t[6854] := 0;
   t[6855] := 0;
   t[6856] := 0;
   t[6857] := 0;
   t[6858] := 0;
   t[6859] := 0;
   t[6860] := 0;
   t[6861] := 0;
   t[6862] := 0;
   t[6863] := 0;
   t[6864] := 0;
   t[6865] := 0;
   t[6866] := 0;
   t[6867] := 0;
   t[6868] := 0;
   t[6869] := 0;
   t[6870] := 0;
   t[6871] := 0;
   t[6872] := 0;
   t[6873] := 0;
   t[6874] := 0;
   t[6875] := 0;
   t[6876] := 0;
   t[6877] := 0;
   t[6878] := 0;
   t[6879] := 0;
   t[6880] := 0;
   t[6881] := 0;
   t[6882] := 0;
   t[6883] := 0;
   t[6884] := 0;
   t[6885] := 0;
   t[6886] := 0;
   t[6887] := 0;
   t[6888] := 0;
   t[6889] := 0;
   t[6890] := 0;
   t[6891] := 0;
   t[6892] := 0;
   t[6893] := 0;
   t[6894] := 0;
   t[6895] := 0;
   t[6896] := 0;
   t[6897] := 0;
   t[6898] := 0;
   t[6899] := 0;
   t[6900] := 0;
   t[6901] := 0;
   t[6902] := 0;
   t[6903] := 0;
   t[6904] := 0;
   t[6905] := 0;
   t[6906] := 0;
   t[6907] := 0;
   t[6908] := 0;
   t[6909] := 0;
   t[6910] := 0;
   t[6911] := 0;
   t[6912] := 0;
   t[6913] := 0;
   t[6914] := 0;
   t[6915] := 0;
   t[6916] := 0;
   t[6917] := 0;
   t[6918] := 0;
   t[6919] := 0;
   t[6920] := 0;
   t[6921] := 0;
   t[6922] := 0;
   t[6923] := 0;
   t[6924] := 0;
   t[6925] := 0;
   t[6926] := 0;
   t[6927] := 0;
   t[6928] := 0;
   t[6929] := 0;
   t[6930] := 0;
   t[6931] := 0;
   t[6932] := 0;
   t[6933] := 0;
   t[6934] := 0;
   t[6935] := 0;
   t[6936] := 0;
   t[6937] := 0;
   t[6938] := 0;
   t[6939] := 0;
   t[6940] := 0;
   t[6941] := 0;
   t[6942] := 0;
   t[6943] := 0;
   t[6944] := 0;
   t[6945] := 0;
   t[6946] := 0;
   t[6947] := 0;
   t[6948] := 0;
   t[6949] := 0;
   t[6950] := 0;
   t[6951] := 0;
   t[6952] := 0;
   t[6953] := 0;
   t[6954] := 0;
   t[6955] := 0;
   t[6956] := 0;
   t[6957] := 0;
   t[6958] := 0;
   t[6959] := 0;
   t[6960] := 0;
   t[6961] := 0;
   t[6962] := 0;
   t[6963] := 0;
   t[6964] := 0;
   t[6965] := 0;
   t[6966] := 0;
   t[6967] := 0;
   t[6968] := 0;
   t[6969] := 0;
   t[6970] := 0;
   t[6971] := 0;
   t[6972] := 0;
   t[6973] := 0;
   t[6974] := 0;
   t[6975] := 0;
   t[6976] := 0;
   t[6977] := 0;
   t[6978] := 0;
   t[6979] := 0;
   t[6980] := 0;
   t[6981] := 0;
   t[6982] := 0;
   t[6983] := 0;
   t[6984] := 0;
   t[6985] := 0;
   t[6986] := 0;
   t[6987] := 0;
   t[6988] := 0;
   t[6989] := 0;
   t[6990] := 0;
   t[6991] := 0;
   t[6992] := 0;
   t[6993] := 0;
   t[6994] := 0;
   t[6995] := 0;
   t[6996] := 0;
   t[6997] := 0;
   t[6998] := 0;
   t[6999] := 0;
   t[7000] := 0;
   t[7001] := 0;
   t[7002] := 0;
   t[7003] := 0;
   t[7004] := 0;
   t[7005] := 0;
   t[7006] := 0;
   t[7007] := 0;
   t[7008] := 0;
   t[7009] := 0;
   t[7010] := 0;
   t[7011] := 0;
   t[7012] := 0;
   t[7013] := 0;
   t[7014] := 0;
   t[7015] := 0;
   t[7016] := 0;
   t[7017] := 0;
   t[7018] := 0;